// TIA Portal project "Street Light Control Based on Light Intensity" (V18)

(* hardware
DEVICE "S7-1200 station_1"  S7-1200 Station
   slot 0: "Rack_0"  S7-1200 Rack  Rack  V1.0
   slot 1: "PLC_1"  CPU 1212C DC/DC/Rly  6ES7 212-1HE40-0XB0  V4.6
DEVICE "HMI_1"  TP900 Comfort
   slot 0: "HMI_1"  TP900 Comfort  6AV2 124-0JC01-0AX0  17.0.0.0
   slot 1: "HMI_RT_1"  TP900 Comfort  6AV2 124-0JC01-0AX0  17.0.0.0
   slot 5: "HMI_1.IE_CP_1"  PROFINET Interface  17.0.0.0
      slot 1: "PROFINET Interface_1"  PROFINET Interface
         slot 1: "Port_1"  Port
         slot 2: "Port_2"  Port
   slot 7: "HMI_1.MPI/DP_CP_1"  MPI/DP Interface  17.0.0.0
*)

// ===== PLC "PLC_1"  CPU 1212C DC/DC/Rly =====

VAR_GLOBAL   // PLC tag table "Default tag table"
   "start" AT %I0.0 : Bool;
   "stop" AT %I0.1 : Bool;
   "power saving" AT %I0.2 : Bool;
   "PIR_sens1" AT %I0.3 : Bool;
   "PIR_sens2" AT %I0.4 : Bool;
   "PIR_sens3" AT %I0.5 : Bool;
   "PIR_sens4" AT %I0.6 : Bool;
   "lamp1" AT %Q0.0 : Bool;
   "lamp2" AT %Q0.1 : Bool;
   "lamp3" AT %Q0.2 : Bool;
   "lamp4" AT %Q0.3 : Bool;
   "lumen" AT %IW64 : Int;
   "system_on_flag" AT %M0.0 : Bool;
   "PIR_status1" AT %M0.1 : Bool;
   "PIR_status2" AT %M0.2 : Bool;
   "PIR_status3" AT %M0.3 : Bool;
   "PIR_status4" AT %M0.4 : Bool;
   "saving1" AT %M0.5 : Bool;
   "saving2" AT %M0.6 : Bool;
   "saving3" AT %M0.7 : Bool;
   "timer_flag" AT %M1.0 : Bool;
END_VAR

ORGANIZATION_BLOCK "Main"   // OB1, LAD, ProgramCycle
TITLE = "Main Program Sweep (Cycle)"
{ S7_Optimized_Access := 'TRUE' }
VERSION : 0.1
   VAR_INPUT
      Initial_Call : Bool;   // Initial call of this OB
      Remanence : Bool;   // =True, if remanent data are available
   END_VAR
   VAR_TEMP   // added for the SCL form of the ladder/FBD networks
      _w1 : Bool;
   END_VAR
BEGIN

REGION Network 1: Start system
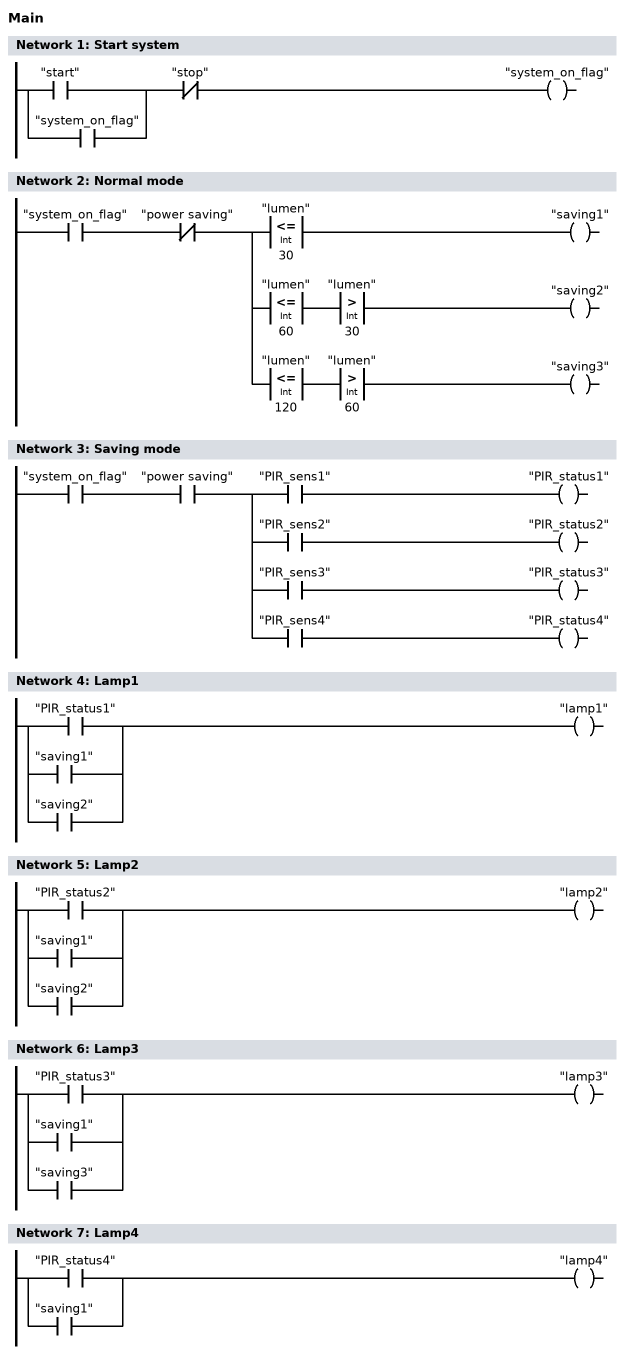
   RUNG wire#powerrail
      Contact( "start" )
      wire#w1
      I_Contact( "stop" )
      Coil( "system_on_flag" )
   END_RUNG
   RUNG wire#powerrail
      Contact( "system_on_flag" )
   END_RUNG wire#w1
   // the same network as SCL:
   "system_on_flag" := ("start" OR "system_on_flag") AND NOT "stop";
END_REGION

REGION Network 2: Normal mode
   RUNG wire#powerrail
      Contact( "system_on_flag" )
      I_Contact( "power saving" )
      wire#w1
      { S7_Templates := "SrcType := Int" } LE_Contact(in1 := "lumen", in2 := 30)
      Coil( "saving1" )
   END_RUNG
   RUNG wire#w1
      { S7_Templates := "SrcType := Int" } LE_Contact(in1 := "lumen", in2 := 60)
      { S7_Templates := "SrcType := Int" } GT_Contact(in1 := "lumen", in2 := 30)
      Coil( "saving2" )
   END_RUNG
   RUNG wire#w1
      { S7_Templates := "SrcType := Int" } LE_Contact(in1 := "lumen", in2 := 120)
      { S7_Templates := "SrcType := Int" } GT_Contact(in1 := "lumen", in2 := 60)
      Coil( "saving3" )
   END_RUNG
   // the same network as SCL:
   #_w1 := "system_on_flag" AND NOT "power saving";
   "saving1" := #_w1 AND ("lumen" <= 30);
   "saving2" := #_w1 AND ("lumen" <= 60) AND ("lumen" > 30);
   "saving3" := #_w1 AND ("lumen" <= 120) AND ("lumen" > 60);
END_REGION

REGION Network 3: Saving mode
   RUNG wire#powerrail
      Contact( "system_on_flag" )
      Contact( "power saving" )
      wire#w1
      Contact( "PIR_sens1" )
      Coil( "PIR_status1" )
   END_RUNG
   RUNG wire#w1
      Contact( "PIR_sens2" )
      Coil( "PIR_status2" )
   END_RUNG
   RUNG wire#w1
      Contact( "PIR_sens3" )
      Coil( "PIR_status3" )
   END_RUNG
   RUNG wire#w1
      Contact( "PIR_sens4" )
      Coil( "PIR_status4" )
   END_RUNG
   // the same network as SCL:
   #_w1 := "system_on_flag" AND "power saving";
   "PIR_status1" := #_w1 AND "PIR_sens1";
   "PIR_status2" := #_w1 AND "PIR_sens2";
   "PIR_status3" := #_w1 AND "PIR_sens3";
   "PIR_status4" := #_w1 AND "PIR_sens4";
END_REGION

REGION Network 4: Lamp1
   RUNG wire#powerrail
      Contact( "PIR_status1" )
      wire#w1
      Coil( "lamp1" )
   END_RUNG
   RUNG wire#powerrail
      Contact( "saving1" )
   END_RUNG wire#w1
   RUNG wire#powerrail
      Contact( "saving2" )
   END_RUNG wire#w1
   // the same network as SCL:
   "lamp1" := "PIR_status1" OR "saving1" OR "saving2";
END_REGION

REGION Network 5: Lamp2
   RUNG wire#powerrail
      Contact( "PIR_status2" )
      wire#w1
      Coil( "lamp2" )
   END_RUNG
   RUNG wire#powerrail
      Contact( "saving1" )
   END_RUNG wire#w1
   RUNG wire#powerrail
      Contact( "saving2" )
   END_RUNG wire#w1
   // the same network as SCL:
   "lamp2" := "PIR_status2" OR "saving1" OR "saving2";
END_REGION

REGION Network 6: Lamp3
   RUNG wire#powerrail
      Contact( "PIR_status3" )
      wire#w1
      Coil( "lamp3" )
   END_RUNG
   RUNG wire#powerrail
      Contact( "saving1" )
   END_RUNG wire#w1
   RUNG wire#powerrail
      Contact( "saving3" )
   END_RUNG wire#w1
   // the same network as SCL:
   "lamp3" := "PIR_status3" OR "saving1" OR "saving3";
END_REGION

REGION Network 7: Lamp4
   RUNG wire#powerrail
      Contact( "PIR_status4" )
      wire#w1
      Coil( "lamp4" )
   END_RUNG
   RUNG wire#powerrail
      Contact( "saving1" )
   END_RUNG wire#w1
   // the same network as SCL:
   "lamp4" := "PIR_status4" OR "saving1";
END_REGION
END_ORGANIZATION_BLOCK

(* ===== HMI "HMI_RT_1" =====
system functions are stored by id; their names below are inferred from use
connection "HMI_Connection_1": ETHERNET, S7_1200_OMS

HMI tags "Default tag table"
   "Lumen" : Int = PLC lumen AT %IW64, 1 s
   "PIR_Sens1" : Bool = PLC PIR_sens1 AT %I0.3, 1 s
   "PIR_Sens2" : Bool = PLC PIR_sens2 AT %I0.4, 1 s
   "PIR_Sens3" : Bool = PLC PIR_sens3 AT %I0.5, 1 s
   "PIR_Sens4" : Bool = PLC PIR_sens4 AT %I0.6, 1 s
   "Lamp1" : Bool = PLC lamp1 AT %Q0.0, 1 s
   "Lamp2" : Bool = PLC lamp2 AT %Q0.1, 1 s
   "Lamp3" : Bool = PLC lamp3 AT %Q0.2, 1 s
   "Lamp4" : Bool = PLC lamp4 AT %Q0.3, 1 s
   "PowerSaving" : Bool = PLC "power saving" AT %I0.2, 1 s
   "Start" : Bool = PLC start AT %I0.0, 1 s
   "Stop" : Bool = PLC stop AT %I0.1, 1 s

Template "Template_1" 800x480
   Button "Exit" at 720,420 size 78x58; TextOff 'Exit'; PictureOff "ExitRuntime_TP900_Comfort_TR"; PictureOn "ExitRuntime_TP900_Comfort_TR"
      on Release: StopRuntime(0)
   Button "Template_Button" at 640,420 size 78x58; TextOff 'Text'
   Button "Template_Button_1" at 560,420 size 78x58; TextOff 'Text'
   Button "Template_Button_2" at 480,420 size 78x58; TextOff 'Text'
   Button "Template_Button_3" at 400,420 size 78x58; TextOff 'Text'
   Button "Template_Button_4" at 321,420 size 78x58; TextOff 'Text'
   Button "Template_Button_5" at 241,420 size 78x58; TextOff 'Text'
   Button "Template_Button_6" at 161,420 size 78x58; TextOff 'Text'
   Button "Alarms" at 81,420 size 78x58; TextOff 'Alarms'; PictureOff "AlarmDisplay_TP900_Comfort_TR"; PictureOn "AlarmDisplay_TP900_Comfort_TR"
      on Release: function_ef3f5d25("Alarm window_Unacknowledged", -1)
   Button "Start screen" at 1,420 size 78x58; TextOff 'Start screen'; PictureOff "NavigateHome_TP900_Comfort_TR"; PictureOn "NavigateHome_TP900_Comfort_TR"
      on Release: ActivateScreen("Root screen", 0)

screen "Root screen" 800x480, template "Template_1"
   GraphicView "Graphic view_1" at 0,2 size 800x418; Picture "IMG_20251103_092201_649(1)(1)"
   Button "Button_2" at 564,181 size 61x40; TextOff 'PIR Sensor 4'
      on Press: function_b14e0dd5("PIR_Sens4", 0)
   Button "Button_3" at 416,181 size 61x40; TextOff 'PIR Sensor 3'
      on Press: function_b14e0dd5("PIR_Sens3", 0)
   Button "Button_4" at 265,181 size 61x40; TextOff 'PIR Sensor 2'
      on Press: function_b14e0dd5("PIR_Sens2", 0)
   Button "Button_5" at 117,181 size 61x40; TextOff 'PIR Sensor 1'
      on Press: function_b14e0dd5("PIR_Sens1", 0)
   Circle "Circle_1" at 496,92 size 20x20
      Visibility <- "Lamp4"
   Circle "Circle_2" at 50,88 size 20x20
      Visibility <- "Lamp1"
   Circle "Circle_3" at 196,92 size 20x20
      Visibility <- "Lamp2"
   Circle "Circle_4" at 349,85 size 22x22
      Visibility <- "Lamp3"
   Switch "Switch_1" at 9,198 size 99x70; CaptionText 'Power Saving'; TextOff 'OFF'; TextOn 'ON'
      ProcessValue <- "PowerSaving"
      on SwitchOn: SetBit("PowerSaving")
      on SwitchOff: ResetBit("PowerSaving")
   Button "Button_6" at 685,287 size 82x43; TextOff 'Start'
      on Press: function_b14e0dd5("Start", 0)
   Button "Button_7" at 30,290 size 82x43; TextOff 'Stop'
      on Press: function_b14e0dd5("Stop", 0)
   IOField "I/O field_1" at 666,88 size 92x51; FormatPattern s99999
      ProcessValue <- "Lumen"
   TextField "Text field_1" at 685,68 size 52x20; Text 'Lumen'
*)